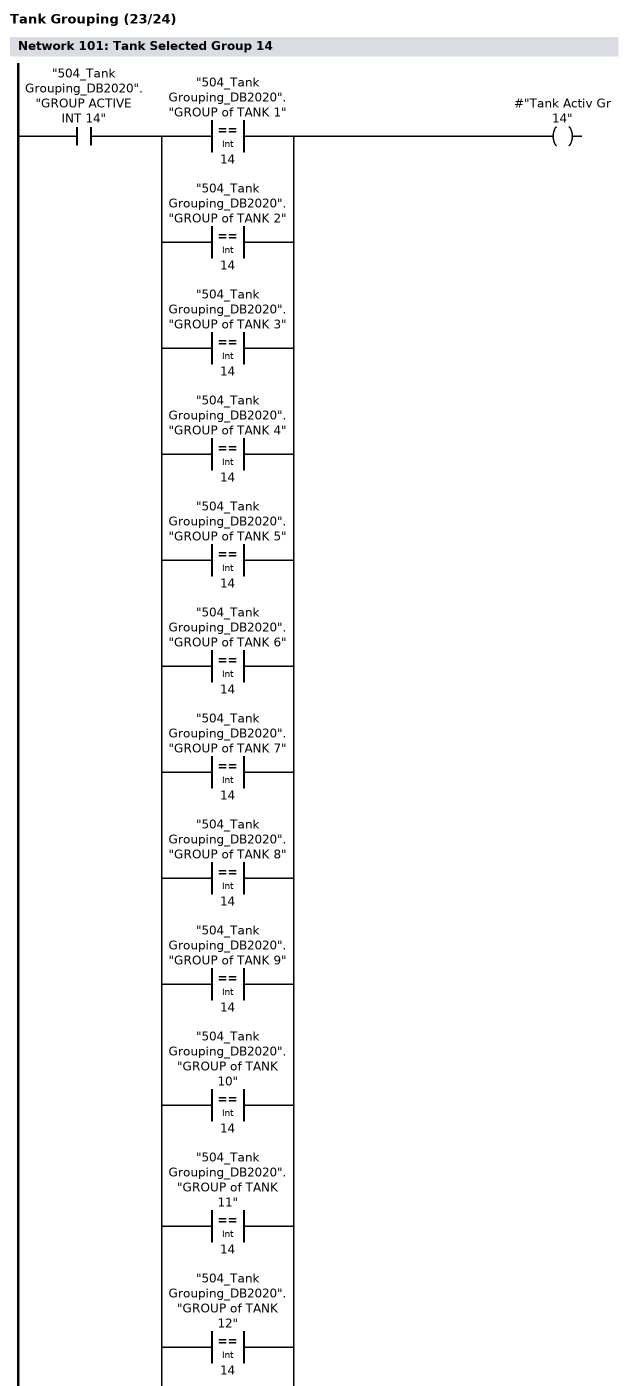
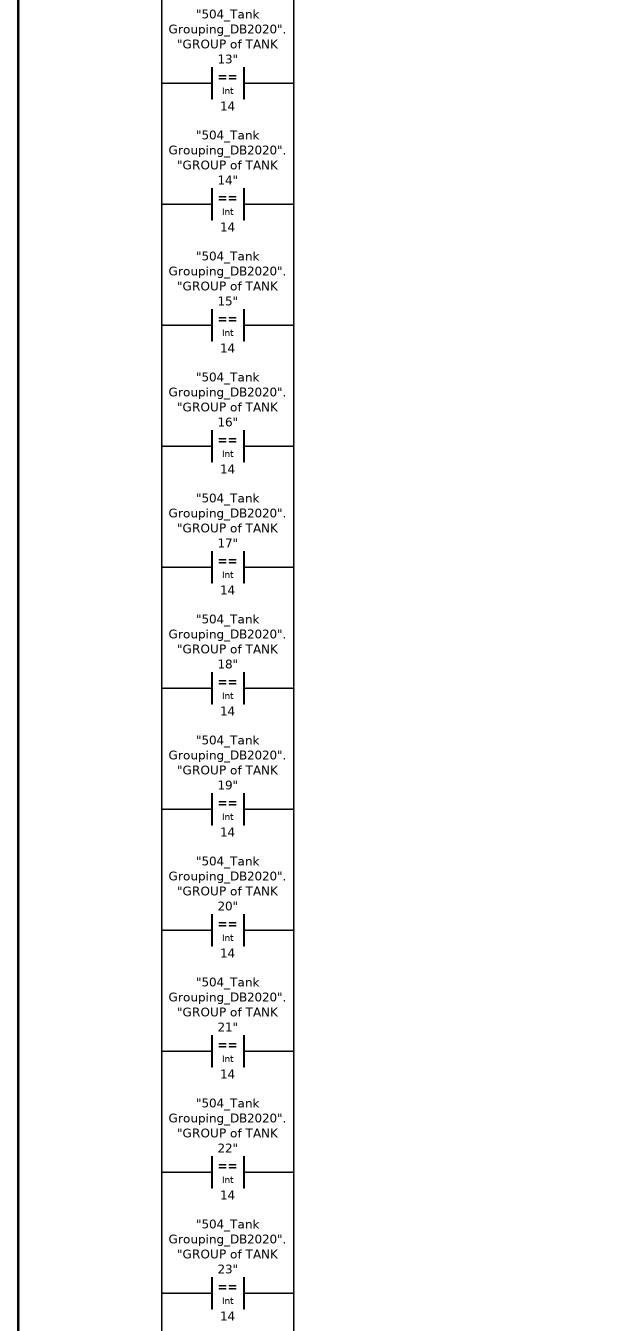
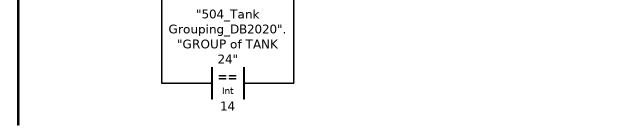
   RUNG wire#powerrail
      Contact( "504_Tank Grouping_DB2020"."GROUP ACTIVE INT 14" )
      wire#w1
      { S7_Templates := "SrcType := Int" } EQ_Contact(in1 := "504_Tank Grouping_DB2020"."GROUP of TANK 1", in2 := 14)
      wire#w2
      Coil( #"Tank Activ Gr 14" )
   END_RUNG
   RUNG wire#w1
      { S7_Templates := "SrcType := Int" } EQ_Contact(in1 := "504_Tank Grouping_DB2020"."GROUP of TANK 2", in2 := 14)
   END_RUNG wire#w2
   RUNG wire#w1
      { S7_Templates := "SrcType := Int" } EQ_Contact(in1 := "504_Tank Grouping_DB2020"."GROUP of TANK 3", in2 := 14)
   END_RUNG wire#w2
   RUNG wire#w1
      { S7_Templates := "SrcType := Int" } EQ_Contact(in1 := "504_Tank Grouping_DB2020"."GROUP of TANK 4", in2 := 14)
   END_RUNG wire#w2
   RUNG wire#w1
      { S7_Templates := "SrcType := Int" } EQ_Contact(in1 := "504_Tank Grouping_DB2020"."GROUP of TANK 5", in2 := 14)
   END_RUNG wire#w2
   RUNG wire#w1
      { S7_Templates := "SrcType := Int" } EQ_Contact(in1 := "504_Tank Grouping_DB2020"."GROUP of TANK 6", in2 := 14)
   END_RUNG wire#w2
   RUNG wire#w1
      { S7_Templates := "SrcType := Int" } EQ_Contact(in1 := "504_Tank Grouping_DB2020"."GROUP of TANK 7", in2 := 14)
   END_RUNG wire#w2
   RUNG wire#w1
      { S7_Templates := "SrcType := Int" } EQ_Contact(in1 := "504_Tank Grouping_DB2020"."GROUP of TANK 8", in2 := 14)
   END_RUNG wire#w2
   RUNG wire#w1
      { S7_Templates := "SrcType := Int" } EQ_Contact(in1 := "504_Tank Grouping_DB2020"."GROUP of TANK 9", in2 := 14)
   END_RUNG wire#w2
   RUNG wire#w1
      { S7_Templates := "SrcType := Int" } EQ_Contact(in1 := "504_Tank Grouping_DB2020"."GROUP of TANK 10", in2 := 14)
   END_RUNG wire#w2
   RUNG wire#w1
      { S7_Templates := "SrcType := Int" } EQ_Contact(in1 := "504_Tank Grouping_DB2020"."GROUP of TANK 11", in2 := 14)
   END_RUNG wire#w2
   RUNG wire#w1
      { S7_Templates := "SrcType := Int" } EQ_Contact(in1 := "504_Tank Grouping_DB2020"."GROUP of TANK 12", in2 := 14)
   END_RUNG wire#w2
   RUNG wire#w1
      { S7_Templates := "SrcType := Int" } EQ_Contact(in1 := "504_Tank Grouping_DB2020"."GROUP of TANK 13", in2 := 14)
   END_RUNG wire#w2
   RUNG wire#w1
      { S7_Templates := "SrcType := Int" } EQ_Contact(in1 := "504_Tank Grouping_DB2020"."GROUP of TANK 14", in2 := 14)
   END_RUNG wire#w2
   RUNG wire#w1
      { S7_Templates := "SrcType := Int" } EQ_Contact(in1 := "504_Tank Grouping_DB2020"."GROUP of TANK 15", in2 := 14)
   END_RUNG wire#w2
   RUNG wire#w1
      { S7_Templates := "SrcType := Int" } EQ_Contact(in1 := "504_Tank Grouping_DB2020"."GROUP of TANK 16", in2 := 14)
   END_RUNG wire#w2
   RUNG wire#w1
      { S7_Templates := "SrcType := Int" } EQ_Contact(in1 := "504_Tank Grouping_DB2020"."GROUP of TANK 17", in2 := 14)
   END_RUNG wire#w2
   RUNG wire#w1
      { S7_Templates := "SrcType := Int" } EQ_Contact(in1 := "504_Tank Grouping_DB2020"."GROUP of TANK 18", in2 := 14)
   END_RUNG wire#w2
   RUNG wire#w1
      { S7_Templates := "SrcType := Int" } EQ_Contact(in1 := "504_Tank Grouping_DB2020"."GROUP of TANK 19", in2 := 14)
   END_RUNG wire#w2
   RUNG wire#w1
      { S7_Templates := "SrcType := Int" } EQ_Contact(in1 := "504_Tank Grouping_DB2020"."GROUP of TANK 20", in2 := 14)
   END_RUNG wire#w2
   RUNG wire#w1
      { S7_Templates := "SrcType := Int" } EQ_Contact(in1 := "504_Tank Grouping_DB2020"."GROUP of TANK 21", in2 := 14)
   END_RUNG wire#w2
   RUNG wire#w1
      { S7_Templates := "SrcType := Int" } EQ_Contact(in1 := "504_Tank Grouping_DB2020"."GROUP of TANK 22", in2 := 14)
   END_RUNG wire#w2
   RUNG wire#w1
      { S7_Templates := "SrcType := Int" } EQ_Contact(in1 := "504_Tank Grouping_DB2020"."GROUP of TANK 23", in2 := 14)
   END_RUNG wire#w2
   RUNG wire#w1
      { S7_Templates := "SrcType := Int" } EQ_Contact(in1 := "504_Tank Grouping_DB2020"."GROUP of TANK 24", in2 := 14)
   END_RUNG wire#w2
   // the same network as SCL:
   #"Tank Activ Gr 14" := "504_Tank Grouping_DB2020"."GROUP ACTIVE INT 14" AND (("504_Tank Grouping_DB2020"."GROUP of TANK 1" = 14) OR ("504_Tank Grouping_DB2020"."GROUP of TANK 2" = 14) OR ("504_Tank Grouping_DB2020"."GROUP of TANK 3" = 14) OR ("504_Tank Grouping_DB2020"."GROUP of TANK 4" = 14) OR ("504_Tank Grouping_DB2020"."GROUP of TANK 5" = 14) OR ("504_Tank Grouping_DB2020"."GROUP of TANK 6" = 14) OR ("504_Tank Grouping_DB2020"."GROUP of TANK 7" = 14) OR ("504_Tank Grouping_DB2020"."GROUP of TANK 8" = 14) OR ("504_Tank Grouping_DB2020"."GROUP of TANK 9" = 14) OR ("504_Tank Grouping_DB2020"."GROUP of TANK 10" = 14) OR ("504_Tank Grouping_DB2020"."GROUP of TANK 11" = 14) OR ("504_Tank Grouping_DB2020"."GROUP of TANK 12" = 14) OR ("504_Tank Grouping_DB2020"."GROUP of TANK 13" = 14) OR ("504_Tank Grouping_DB2020"."GROUP of TANK 14" = 14) OR ("504_Tank Grouping_DB2020"."GROUP of TANK 15" = 14) OR ("504_Tank Grouping_DB2020"."GROUP of TANK 16" = 14) OR ("504_Tank Grouping_DB2020"."GROUP of TANK 17" = 14) OR ("504_Tank Grouping_DB2020"."GROUP of TANK 18" = 14) OR ("504_Tank Grouping_DB2020"."GROUP of TANK 19" = 14) OR ("504_Tank Grouping_DB2020"."GROUP of TANK 20" = 14) OR ("504_Tank Grouping_DB2020"."GROUP of TANK 21" = 14) OR ("504_Tank Grouping_DB2020"."GROUP of TANK 22" = 14) OR ("504_Tank Grouping_DB2020"."GROUP of TANK 23" = 14) OR ("504_Tank Grouping_DB2020"."GROUP of TANK 24" = 14));
END_REGION

REGION Network 102: Tank Selected Group
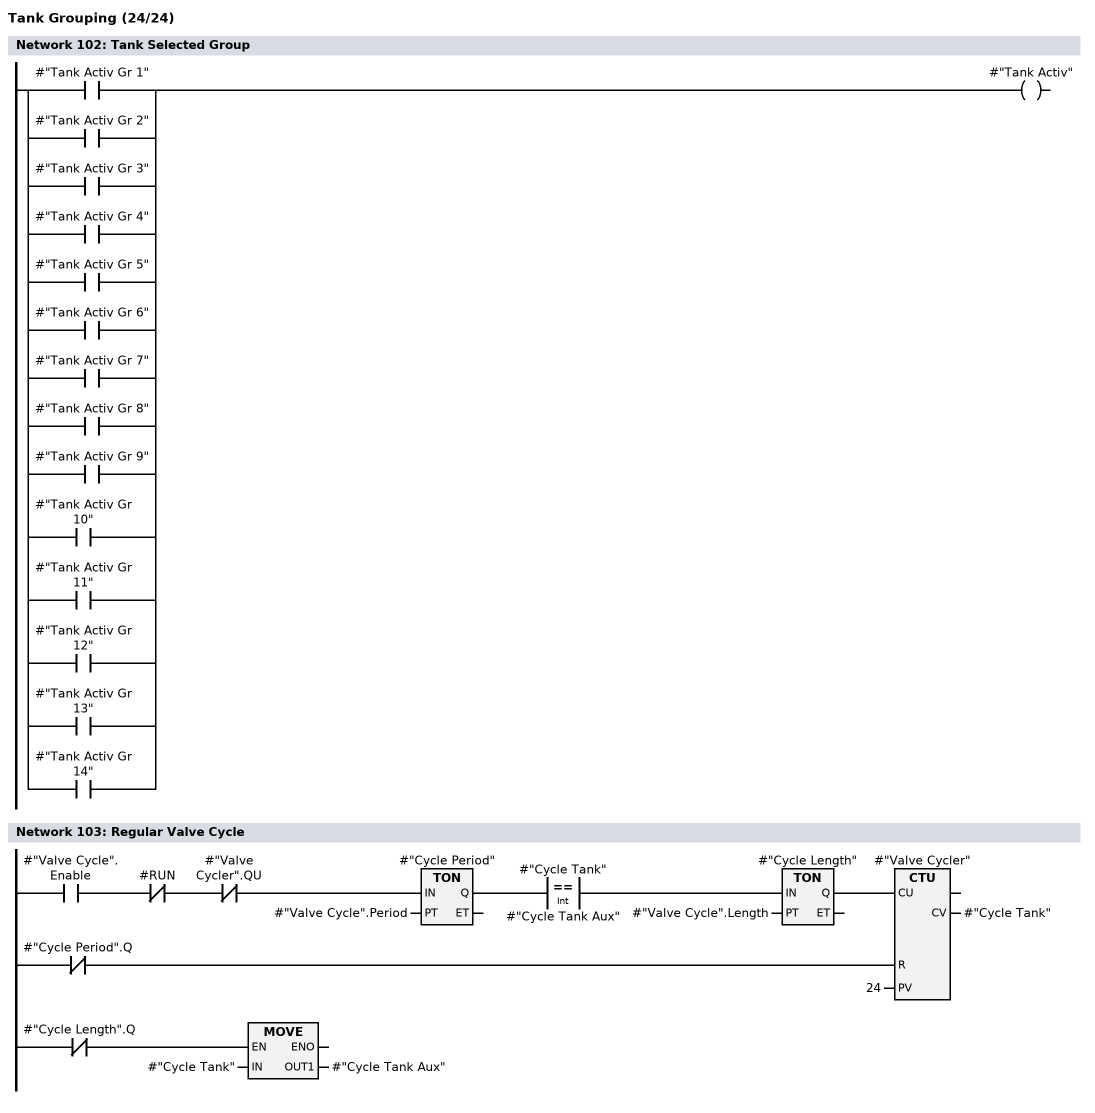
   RUNG wire#powerrail
      Contact( #"Tank Activ Gr 1" )
      wire#w1
      Coil( #"Tank Activ" )
   END_RUNG
   RUNG wire#powerrail
      Contact( #"Tank Activ Gr 2" )
   END_RUNG wire#w1
   RUNG wire#powerrail
      Contact( #"Tank Activ Gr 3" )
   END_RUNG wire#w1
   RUNG wire#powerrail
      Contact( #"Tank Activ Gr 4" )
   END_RUNG wire#w1
   RUNG wire#powerrail
      Contact( #"Tank Activ Gr 5" )
   END_RUNG wire#w1
   RUNG wire#powerrail
      Contact( #"Tank Activ Gr 6" )
   END_RUNG wire#w1
   RUNG wire#powerrail
      Contact( #"Tank Activ Gr 7" )
   END_RUNG wire#w1
   RUNG wire#powerrail
      Contact( #"Tank Activ Gr 8" )
   END_RUNG wire#w1
   RUNG wire#powerrail
      Contact( #"Tank Activ Gr 9" )
   END_RUNG wire#w1
   RUNG wire#powerrail
      Contact( #"Tank Activ Gr 10" )
   END_RUNG wire#w1
   RUNG wire#powerrail
      Contact( #"Tank Activ Gr 11" )
   END_RUNG wire#w1
   RUNG wire#powerrail
      Contact( #"Tank Activ Gr 12" )
   END_RUNG wire#w1
   RUNG wire#powerrail
      Contact( #"Tank Activ Gr 13" )
   END_RUNG wire#w1
   RUNG wire#powerrail
      Contact( #"Tank Activ Gr 14" )
   END_RUNG wire#w1
   // the same network as SCL:
   #"Tank Activ" := #"Tank Activ Gr 1" OR #"Tank Activ Gr 2" OR #"Tank Activ Gr 3" OR #"Tank Activ Gr 4" OR #"Tank Activ Gr 5" OR #"Tank Activ Gr 6" OR #"Tank Activ Gr 7" OR #"Tank Activ Gr 8" OR #"Tank Activ Gr 9" OR #"Tank Activ Gr 10" OR #"Tank Activ Gr 11" OR #"Tank Activ Gr 12" OR #"Tank Activ Gr 13" OR #"Tank Activ Gr 14";
END_REGION

REGION Network 103: Regular Valve Cycle
   #"Cycle Period"(IN := #"Valve Cycle".Enable AND NOT #RUN AND NOT #"Valve Cycler".QU,   // TON
                   PT := #"Valve Cycle".Period);
   #"Cycle Length"(IN := #"Cycle Period".Q AND (#"Cycle Tank" = #"Cycle Tank Aux"), PT := #"Valve Cycle".Length);   // TON
   #"Valve Cycler"(CU := #"Cycle Length".Q, R := NOT #"Cycle Period".Q, PV := 24, CV => #"Cycle Tank");   // CTU
   IF NOT #"Cycle Length".Q THEN #"Cycle Tank Aux" := #"Cycle Tank"; END_IF;
END_REGION
END_FUNCTION_BLOCK

FUNCTION_BLOCK "505_GROUP SEQUENCE"   // FB505, LAD
{ S7_Optimized_Access := 'TRUE' }
VERSION : 0.1
   VAR_INPUT
      Run : Bool;
      "Sequence Time Min" : Int;
      "Setpoint Time Min" : Int;
      "Sequence Time Min Delay" : Int;
      "O2 Confirmed Time" : Int;
      "RIO 1" : "3T_IP_DATA";
      "RIO 2" : "2T_IP_DATA";
      "RIO 3" : "2T_IP_DATA";
      "RIO 4" : "2T_IP_DATA";
      "RIO 5" : "2T_IP_DATA";
      "RIO 6" : "2T_IP_DATA";
      "RIO 7" : "1T_IP_DATA";
      "GROUP ACTIV 1" : Bool;
      "GROUP ACTIV 2" : Bool;
      "GROUP ACTIV 3" : Bool;
      "GROUP ACTIV 4" : Bool;
      "GROUP ACTIV 5" : Bool;
      "GROUP ACTIV 6" : Bool;
      "GROUP ACTIV 7" : Bool;
      "1Hz" : Bool;
   END_VAR
   VAR_OUTPUT
      "Sequence Time Min Remaining_Reset" : Int;
      "Setpoint Time Min Remaining_Reset" : Int;
      "RUN GROUP 1" : Bool;
      "RUN GROUP 2" : Bool;
      "RUN GROUP 3" : Bool;
      "RUN GROUP 4" : Bool;
      "RUN GROUP 5" : Bool;
      "RUN GROUP 6" : Bool;
      "RUN GROUP 7" : Bool;
   END_VAR
   VAR
      "1Hz Puls" : Bool;
      "1Hz Puls_Aux" : Bool;
      "Sequence Time Min Remaining G 1" : Int;
      "Sequence Time Min Remaining G 2" : Int;
      "Sequence Time Min Remaining G 3" : Int;
      "Sequence Time Min Remaining G 4" : Int;
      "Sequence Time Min Remaining G 5" : Int;
      "Sequence Time Min Remaining G 6" : Int;
      "Sequence Time Min Remaining G 7" : Int;
      "Sequence Time Min Delay G 1" : Int;
      "Sequence Time Min Delay G 2" : Int;
      "Sequence Time Min Delay G 3" : Int;
      "Sequence Time Min Delay G 4" : Int;
      "Sequence Time Min Delay G 5" : Int;
      "Sequence Time Min Delay G 6" : Int;
      "Sequence Time Min Delay G 7" : Int;
      "Setpoint Time Min Remaining G 1" : Int;
      "Setpoint Time Min Remaining G 2" : Int;
      "Setpoint Time Min Remaining G 3" : Int;
      "Setpoint Time Min Remaining G 4" : Int;
      "Setpoint Time Min Remaining G 5" : Int;
      "Setpoint Time Min Remaining G 6" : Int;
      "Setpoint Time Min Remaining G 7" : Int;
      Second : Int;
      Minut : Int;
      Minut_Puls : Bool;
      R_TRIG_Instance : R_TRIG;
      Aux : Struct
         "Aux 1" : Bool;
         "Aux 2" : Bool;
         "Aux 3" : Bool;
         "Aux 4" : Bool;
         "Aux 5" : Bool;
         "Aux 6" : Bool;
         "Aux 7" : Bool;
      END_STRUCT;
   END_VAR
   VAR_TEMP   // added for the SCL form of the ladder/FBD networks
      _w1 : Bool;
      _w2 : Bool;
   END_VAR
BEGIN

REGION Network 1: 1Hz Puls
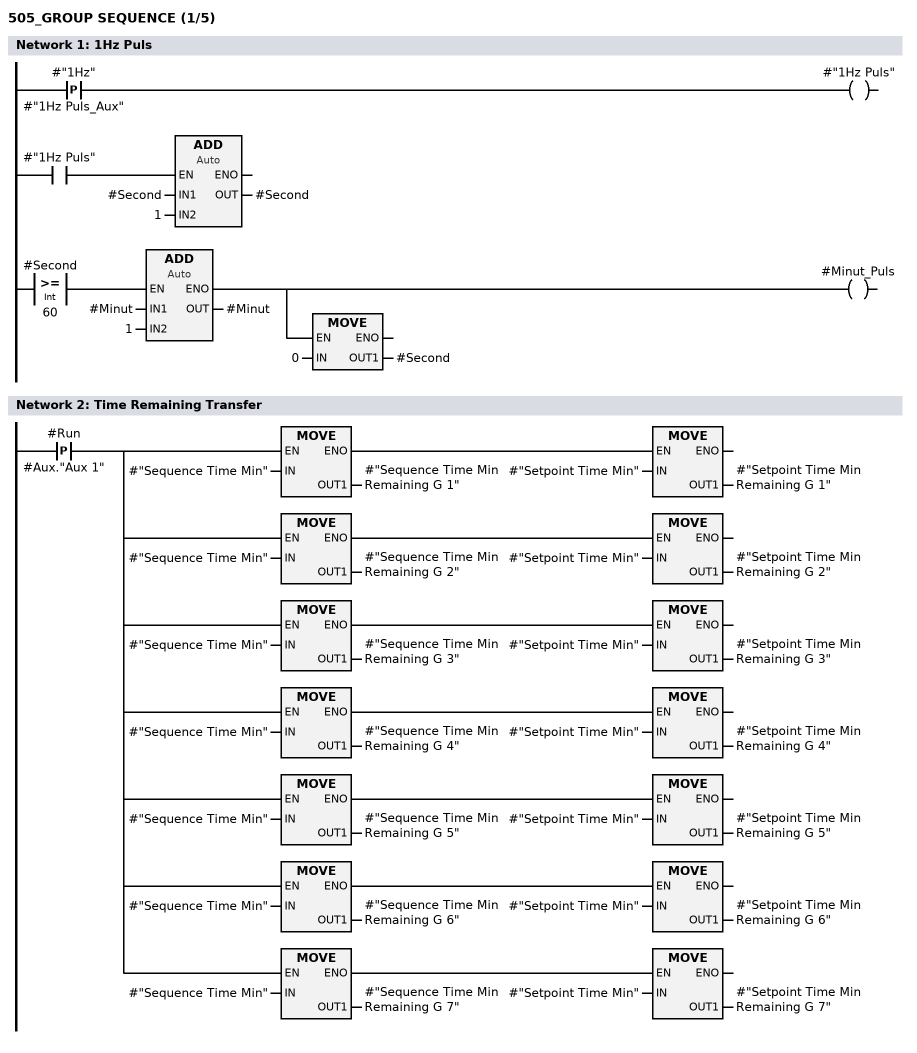
   RUNG wire#powerrail
      P_Contact(operand := #"1Hz", bit := #"1Hz Puls_Aux")
      Coil( #"1Hz Puls" )
   END_RUNG
   RUNG wire#powerrail
      Contact( #"1Hz Puls" )
      Add(in1 := #Second, in2 := 1, out => #Second)
   END_RUNG
   RUNG wire#powerrail
      { S7_Templates := "SrcType := Int" } GE_Contact(in1 := #Second, in2 := 60)
      Add(in1 := #Minut, in2 := 1, out => #Minut)
      wire#w1
      Coil( #Minut_Puls )
   END_RUNG
   RUNG wire#w1
      Move(in := 0, out1 => #Second)
   END_RUNG
   // the same network as SCL:
   #_w1 := #"1Hz" AND NOT #"1Hz Puls_Aux";   // rising edge of #"1Hz"
   #"1Hz Puls_Aux" := #"1Hz";
   #"1Hz Puls" := #_w1;
   IF #"1Hz Puls" THEN #Second := #Second + 1; END_IF;
   #_w2 := #Second >= 60;
   IF #_w2 THEN #Minut := #Minut + 1; END_IF;
   #Minut_Puls := #_w2;
   IF #_w2 THEN #Second := 0; END_IF;
END_REGION

REGION Network 2: Time Remaining Transfer
   RUNG wire#powerrail
      P_Contact(operand := #Run, bit := #Aux."Aux 1")
      wire#w1
      Move(in := #"Sequence Time Min", out1 => #"Sequence Time Min Remaining G 1")
      Move(in := #"Setpoint Time Min", out1 => #"Setpoint Time Min Remaining G 1")
   END_RUNG
   RUNG wire#w1
      Move(in := #"Sequence Time Min", out1 => #"Sequence Time Min Remaining G 2")
      Move(in := #"Setpoint Time Min", out1 => #"Setpoint Time Min Remaining G 2")
   END_RUNG
   RUNG wire#w1
      Move(in := #"Sequence Time Min", out1 => #"Sequence Time Min Remaining G 3")
      Move(in := #"Setpoint Time Min", out1 => #"Setpoint Time Min Remaining G 3")
   END_RUNG
   RUNG wire#w1
      Move(in := #"Sequence Time Min", out1 => #"Sequence Time Min Remaining G 4")
      Move(in := #"Setpoint Time Min", out1 => #"Setpoint Time Min Remaining G 4")
   END_RUNG
   RUNG wire#w1
      Move(in := #"Sequence Time Min", out1 => #"Sequence Time Min Remaining G 5")
      Move(in := #"Setpoint Time Min", out1 => #"Setpoint Time Min Remaining G 5")
   END_RUNG
   RUNG wire#w1
      Move(in := #"Sequence Time Min", out1 => #"Sequence Time Min Remaining G 6")
      Move(in := #"Setpoint Time Min", out1 => #"Setpoint Time Min Remaining G 6")
   END_RUNG
   RUNG wire#w1
      Move(in := #"Sequence Time Min", out1 => #"Sequence Time Min Remaining G 7")
      Move(in := #"Setpoint Time Min", out1 => #"Setpoint Time Min Remaining G 7")
   END_RUNG
   // the same network as SCL:
   #_w1 := #Run AND NOT #Aux."Aux 1";   // rising edge of #Run
   #Aux."Aux 1" := #Run;
   IF #_w1 THEN
       #"Sequence Time Min Remaining G 1" := #"Sequence Time Min";
       #"Setpoint Time Min Remaining G 1" := #"Setpoint Time Min";
       #"Sequence Time Min Remaining G 2" := #"Sequence Time Min";
       #"Setpoint Time Min Remaining G 2" := #"Setpoint Time Min";
       #"Sequence Time Min Remaining G 3" := #"Sequence Time Min";
       #"Setpoint Time Min Remaining G 3" := #"Setpoint Time Min";
       #"Sequence Time Min Remaining G 4" := #"Sequence Time Min";
       #"Setpoint Time Min Remaining G 4" := #"Setpoint Time Min";
       #"Sequence Time Min Remaining G 5" := #"Sequence Time Min";
       #"Setpoint Time Min Remaining G 5" := #"Setpoint Time Min";
       #"Sequence Time Min Remaining G 6" := #"Sequence Time Min";
       #"Setpoint Time Min Remaining G 6" := #"Setpoint Time Min";
       #"Sequence Time Min Remaining G 7" := #"Sequence Time Min";
       #"Setpoint Time Min Remaining G 7" := #"Setpoint Time Min";
   END_IF;
END_REGION

REGION Network 3: Delay Transfer
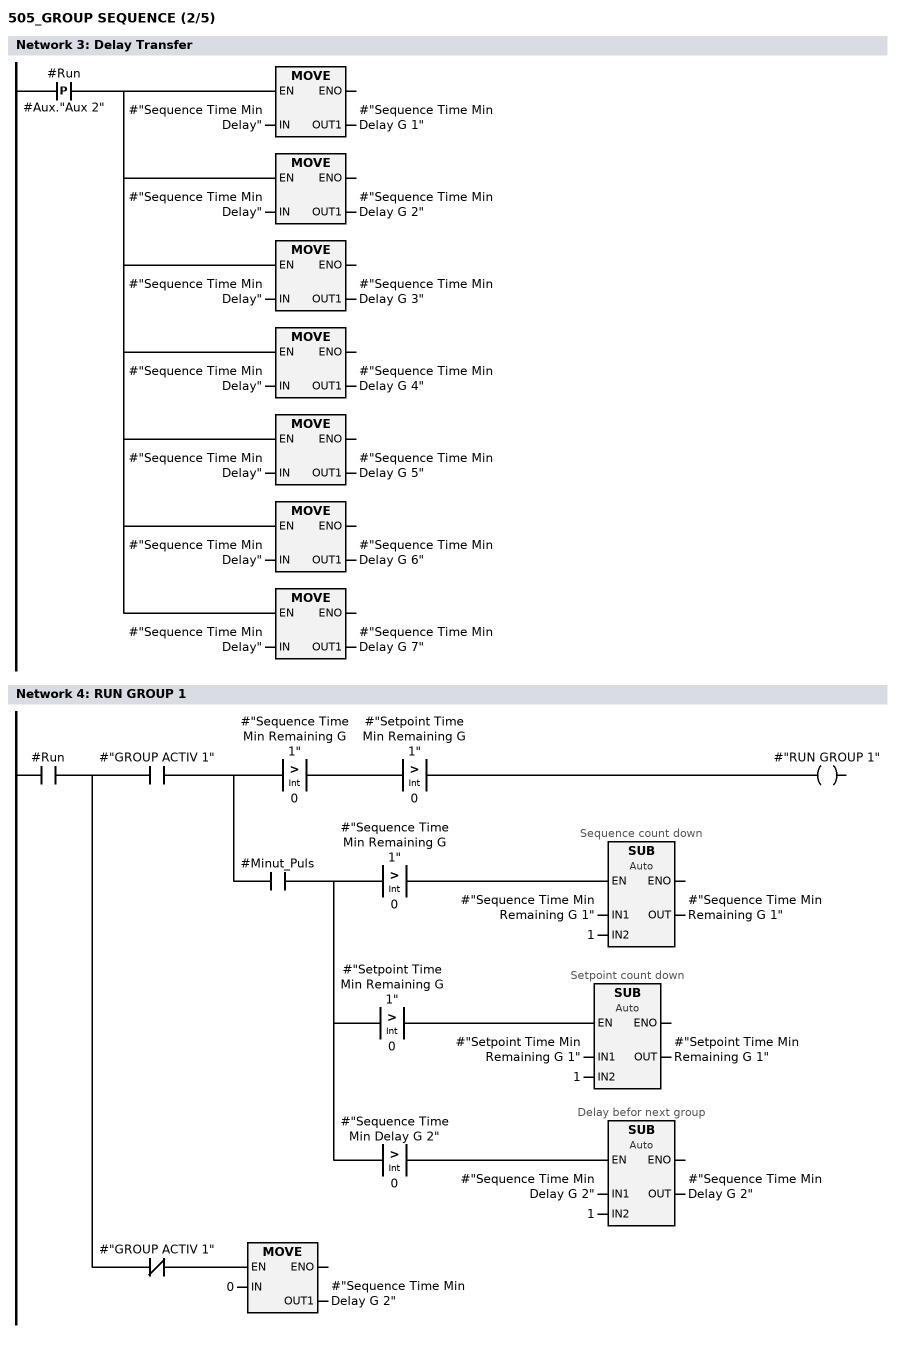
   RUNG wire#powerrail
      P_Contact(operand := #Run, bit := #Aux."Aux 2")
      wire#w1
      Move(in := #"Sequence Time Min Delay", out1 => #"Sequence Time Min Delay G 1")
   END_RUNG
   RUNG wire#w1
      Move(in := #"Sequence Time Min Delay", out1 => #"Sequence Time Min Delay G 2")
   END_RUNG
   RUNG wire#w1
      Move(in := #"Sequence Time Min Delay", out1 => #"Sequence Time Min Delay G 3")
   END_RUNG
   RUNG wire#w1
      Move(in := #"Sequence Time Min Delay", out1 => #"Sequence Time Min Delay G 4")
   END_RUNG
   RUNG wire#w1
      Move(in := #"Sequence Time Min Delay", out1 => #"Sequence Time Min Delay G 5")
   END_RUNG
   RUNG wire#w1
      Move(in := #"Sequence Time Min Delay", out1 => #"Sequence Time Min Delay G 6")
   END_RUNG
   RUNG wire#w1
      Move(in := #"Sequence Time Min Delay", out1 => #"Sequence Time Min Delay G 7")
   END_RUNG
   // the same network as SCL:
   #_w1 := #Run AND NOT #Aux."Aux 2";   // rising edge of #Run
   #Aux."Aux 2" := #Run;
   IF #_w1 THEN
       #"Sequence Time Min Delay G 1" := #"Sequence Time Min Delay";
       #"Sequence Time Min Delay G 2" := #"Sequence Time Min Delay";
       #"Sequence Time Min Delay G 3" := #"Sequence Time Min Delay";
       #"Sequence Time Min Delay G 4" := #"Sequence Time Min Delay";
       #"Sequence Time Min Delay G 5" := #"Sequence Time Min Delay";
       #"Sequence Time Min Delay G 6" := #"Sequence Time Min Delay";
       #"Sequence Time Min Delay G 7" := #"Sequence Time Min Delay";
   END_IF;
END_REGION

REGION Network 4: RUN GROUP 1
   RUNG wire#powerrail
      Contact( #Run )
      wire#w1
      Contact( #"GROUP ACTIV 1" )
      wire#w2
      { S7_Templates := "SrcType := Int" } GT_Contact(in1 := #"Sequence Time Min Remaining G 1", in2 := 0)
      { S7_Templates := "SrcType := Int" } GT_Contact(in1 := #"Setpoint Time Min Remaining G 1", in2 := 0)
      Coil( #"RUN GROUP 1" )
   END_RUNG
   RUNG wire#w2
      Contact( #Minut_Puls )
      wire#w3
      { S7_Templates := "SrcType := Int" } GT_Contact(in1 := #"Sequence Time Min Remaining G 1", in2 := 0)
      Sub(in1 := #"Sequence Time Min Remaining G 1", in2 := 1, out => #"Sequence Time Min Remaining G 1")   // Sequence count down
   END_RUNG
   RUNG wire#w3
      { S7_Templates := "SrcType := Int" } GT_Contact(in1 := #"Setpoint Time Min Remaining G 1", in2 := 0)
      Sub(in1 := #"Setpoint Time Min Remaining G 1", in2 := 1, out => #"Setpoint Time Min Remaining G 1")   // Setpoint count down
   END_RUNG
   RUNG wire#w3
      { S7_Templates := "SrcType := Int" } GT_Contact(in1 := #"Sequence Time Min Delay G 2", in2 := 0)
      Sub(in1 := #"Sequence Time Min Delay G 2", in2 := 1, out => #"Sequence Time Min Delay G 2")   // Delay befor next group
   END_RUNG
   RUNG wire#w1
      I_Contact( #"GROUP ACTIV 1" )
      Move(in := 0, out1 => #"Sequence Time Min Delay G 2")
   END_RUNG
   // the same network as SCL:
   #_w1 := #Run AND #"GROUP ACTIV 1";
   #"RUN GROUP 1" := #_w1 AND (#"Sequence Time Min Remaining G 1" > 0) AND (#"Setpoint Time Min Remaining G 1" > 0);
   #_w2 := #_w1 AND #Minut_Puls;
   IF #_w2 AND (#"Sequence Time Min Remaining G 1" > 0) THEN
       #"Sequence Time Min Remaining G 1" := #"Sequence Time Min Remaining G 1" - 1;   // Sequence count down
   END_IF;
   IF #_w2 AND (#"Setpoint Time Min Remaining G 1" > 0) THEN
       #"Setpoint Time Min Remaining G 1" := #"Setpoint Time Min Remaining G 1" - 1;   // Setpoint count down
   END_IF;
   IF #_w2 AND (#"Sequence Time Min Delay G 2" > 0) THEN
       #"Sequence Time Min Delay G 2" := #"Sequence Time Min Delay G 2" - 1;   // Delay befor next group
   END_IF;
   IF #Run AND NOT #"GROUP ACTIV 1" THEN #"Sequence Time Min Delay G 2" := 0; END_IF;
END_REGION

REGION Network 5: RUN GROUP 2
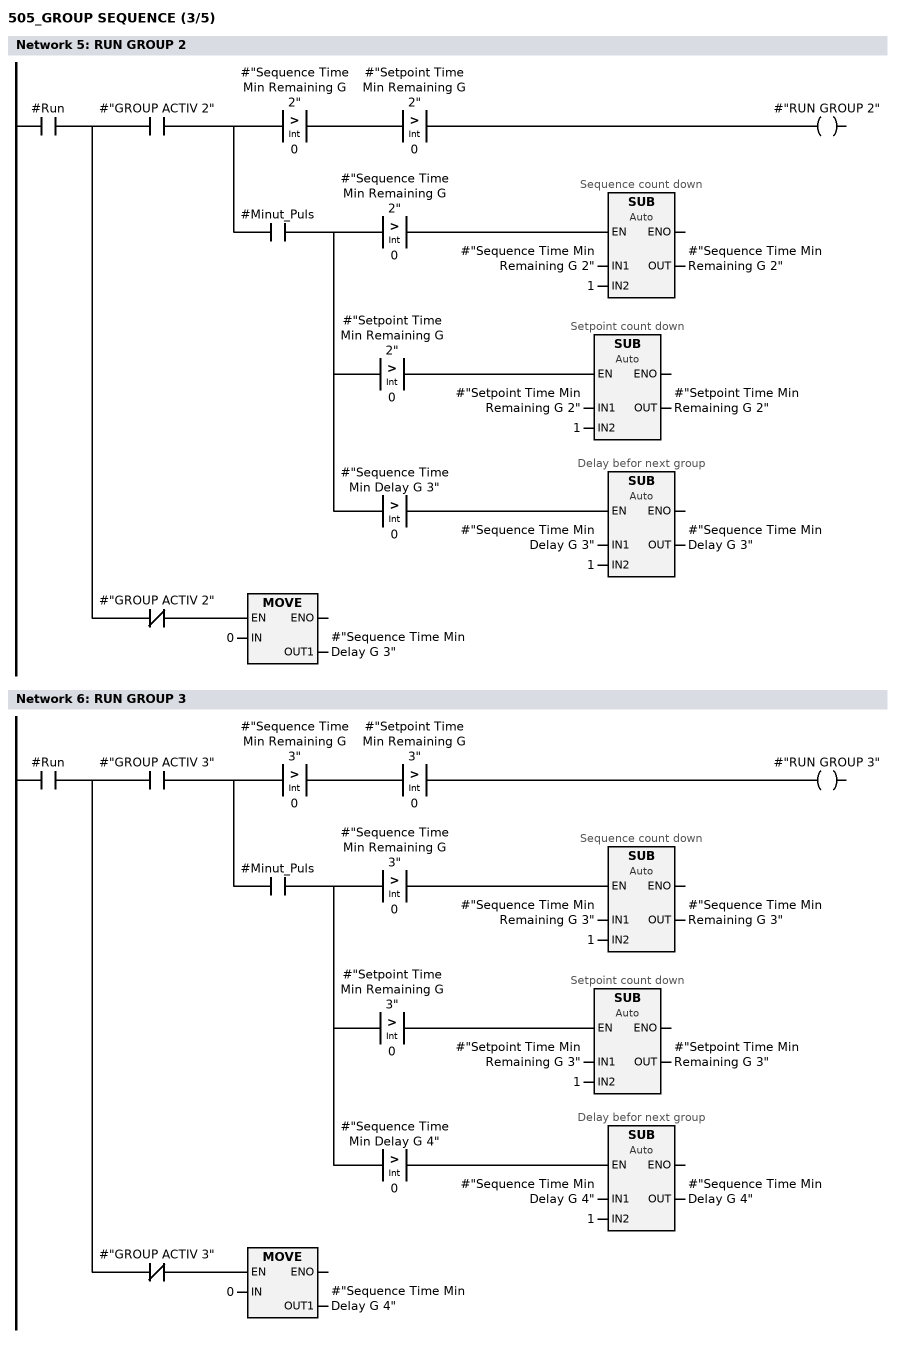
   RUNG wire#powerrail
      Contact( #Run )
      wire#w1
      Contact( #"GROUP ACTIV 2" )
      wire#w2
      { S7_Templates := "SrcType := Int" } GT_Contact(in1 := #"Sequence Time Min Remaining G 2", in2 := 0)
      { S7_Templates := "SrcType := Int" } GT_Contact(in1 := #"Setpoint Time Min Remaining G 2", in2 := 0)
      Coil( #"RUN GROUP 2" )
   END_RUNG
   RUNG wire#w2
      Contact( #Minut_Puls )
      wire#w3
      { S7_Templates := "SrcType := Int" } GT_Contact(in1 := #"Sequence Time Min Remaining G 2", in2 := 0)
      Sub(in1 := #"Sequence Time Min Remaining G 2", in2 := 1, out => #"Sequence Time Min Remaining G 2")   // Sequence count down
   END_RUNG
   RUNG wire#w3
      { S7_Templates := "SrcType := Int" } GT_Contact(in1 := #"Setpoint Time Min Remaining G 2", in2 := 0)
      Sub(in1 := #"Setpoint Time Min Remaining G 2", in2 := 1, out => #"Setpoint Time Min Remaining G 2")   // Setpoint count down
   END_RUNG
   RUNG wire#w3
      { S7_Templates := "SrcType := Int" } GT_Contact(in1 := #"Sequence Time Min Delay G 3", in2 := 0)
      Sub(in1 := #"Sequence Time Min Delay G 3", in2 := 1, out => #"Sequence Time Min Delay G 3")   // Delay befor next group
   END_RUNG
   RUNG wire#w1
      I_Contact( #"GROUP ACTIV 2" )
      Move(in := 0, out1 => #"Sequence Time Min Delay G 3")
   END_RUNG
   // the same network as SCL:
   #_w1 := #Run AND #"GROUP ACTIV 2";
   #"RUN GROUP 2" := #_w1 AND (#"Sequence Time Min Remaining G 2" > 0) AND (#"Setpoint Time Min Remaining G 2" > 0);
   #_w2 := #_w1 AND #Minut_Puls;
   IF #_w2 AND (#"Sequence Time Min Remaining G 2" > 0) THEN
       #"Sequence Time Min Remaining G 2" := #"Sequence Time Min Remaining G 2" - 1;   // Sequence count down
   END_IF;
   IF #_w2 AND (#"Setpoint Time Min Remaining G 2" > 0) THEN
       #"Setpoint Time Min Remaining G 2" := #"Setpoint Time Min Remaining G 2" - 1;   // Setpoint count down
   END_IF;
   IF #_w2 AND (#"Sequence Time Min Delay G 3" > 0) THEN
       #"Sequence Time Min Delay G 3" := #"Sequence Time Min Delay G 3" - 1;   // Delay befor next group
   END_IF;
   IF #Run AND NOT #"GROUP ACTIV 2" THEN #"Sequence Time Min Delay G 3" := 0; END_IF;
END_REGION

REGION Network 6: RUN GROUP 3
   RUNG wire#powerrail
      Contact( #Run )
      wire#w1
      Contact( #"GROUP ACTIV 3" )
      wire#w2
      { S7_Templates := "SrcType := Int" } GT_Contact(in1 := #"Sequence Time Min Remaining G 3", in2 := 0)
      { S7_Templates := "SrcType := Int" } GT_Contact(in1 := #"Setpoint Time Min Remaining G 3", in2 := 0)
      Coil( #"RUN GROUP 3" )
   END_RUNG
   RUNG wire#w2
      Contact( #Minut_Puls )
      wire#w3
      { S7_Templates := "SrcType := Int" } GT_Contact(in1 := #"Sequence Time Min Remaining G 3", in2 := 0)
      Sub(in1 := #"Sequence Time Min Remaining G 3", in2 := 1, out => #"Sequence Time Min Remaining G 3")   // Sequence count down
   END_RUNG
   RUNG wire#w3
      { S7_Templates := "SrcType := Int" } GT_Contact(in1 := #"Setpoint Time Min Remaining G 3", in2 := 0)
      Sub(in1 := #"Setpoint Time Min Remaining G 3", in2 := 1, out => #"Setpoint Time Min Remaining G 3")   // Setpoint count down
   END_RUNG
   RUNG wire#w3
      { S7_Templates := "SrcType := Int" } GT_Contact(in1 := #"Sequence Time Min Delay G 4", in2 := 0)
      Sub(in1 := #"Sequence Time Min Delay G 4", in2 := 1, out => #"Sequence Time Min Delay G 4")   // Delay befor next group
   END_RUNG
   RUNG wire#w1
      I_Contact( #"GROUP ACTIV 3" )
      Move(in := 0, out1 => #"Sequence Time Min Delay G 4")
   END_RUNG
   // the same network as SCL:
   #_w1 := #Run AND #"GROUP ACTIV 3";
   #"RUN GROUP 3" := #_w1 AND (#"Sequence Time Min Remaining G 3" > 0) AND (#"Setpoint Time Min Remaining G 3" > 0);
   #_w2 := #_w1 AND #Minut_Puls;
   IF #_w2 AND (#"Sequence Time Min Remaining G 3" > 0) THEN
       #"Sequence Time Min Remaining G 3" := #"Sequence Time Min Remaining G 3" - 1;   // Sequence count down
   END_IF;
   IF #_w2 AND (#"Setpoint Time Min Remaining G 3" > 0) THEN
       #"Setpoint Time Min Remaining G 3" := #"Setpoint Time Min Remaining G 3" - 1;   // Setpoint count down
   END_IF;
   IF #_w2 AND (#"Sequence Time Min Delay G 4" > 0) THEN
       #"Sequence Time Min Delay G 4" := #"Sequence Time Min Delay G 4" - 1;   // Delay befor next group
   END_IF;
   IF #Run AND NOT #"GROUP ACTIV 3" THEN #"Sequence Time Min Delay G 4" := 0; END_IF;
END_REGION

REGION Network 7: RUN GROUP 4